(* Logix 5000 project; controller OWF Emulate 5570 rev 30.12; software revision 30.00 *) (continued)
   	OWF_Key[222,1]:=1243582292;
   	OWF_Key[222,2]:=1667078718;
   	OWF_Key[222,3]:=820047921;
   	OWF_Key[222,4]:=2100818839;
   	OWF_Key[222,5]:=54664303;
   	OWF_Key[222,6]:=832390246;
   	OWF_Key[222,7]:=1025838178;
   	OWF_Key[222,8]:=2108609866;
   	OWF_Key[223,0]:=1550121582;
   	OWF_Key[223,1]:=901840231;
   	OWF_Key[223,2]:=845237975;
   	OWF_Key[223,3]:=1737038115;
   	OWF_Key[223,4]:=250371253;
   	OWF_Key[223,5]:=841400060;
   	OWF_Key[223,6]:=633458828;
   	OWF_Key[223,7]:=1234192716;
   	OWF_Key[223,8]:=1638825880;
   	OWF_Key[224,0]:=1100202784;
   	OWF_Key[224,1]:=1268618722;
   	OWF_Key[224,2]:=1328247563;
   	OWF_Key[224,3]:=315030373;
   	OWF_Key[224,4]:=17465755;
   	OWF_Key[224,5]:=1489898403;
   	OWF_Key[224,6]:=1369322265;
   	OWF_Key[224,7]:=2029664960;
   	OWF_Key[224,8]:=1183192871;
   	OWF_Key[225,0]:=1841076227;
   	OWF_Key[225,1]:=1387440943;
   	OWF_Key[225,2]:=94964990;
   	OWF_Key[225,3]:=374620338;
   	OWF_Key[225,4]:=198656364;
   	OWF_Key[225,5]:=451329169;
   	OWF_Key[225,6]:=1040984125;
   	OWF_Key[225,7]:=421870535;
   	OWF_Key[225,8]:=1711294224;
   	OWF_Key[226,0]:=908174588;
   	OWF_Key[226,1]:=915800259;
   	OWF_Key[226,2]:=1938292132;
   	OWF_Key[226,3]:=1295597437;
   	OWF_Key[226,4]:=543239841;
   	OWF_Key[226,5]:=543313500;
   	OWF_Key[226,6]:=1320318736;
   	OWF_Key[226,7]:=1310833438;
   	OWF_Key[226,8]:=1604355088;
   	OWF_Key[227,0]:=1963899269;
   	OWF_Key[227,1]:=1680451206;
   	OWF_Key[227,2]:=236776837;
   	OWF_Key[227,3]:=1960573892;
   	OWF_Key[227,4]:=2100303206;
   	OWF_Key[227,5]:=407078522;
   	OWF_Key[227,6]:=949933681;
   	OWF_Key[227,7]:=279399557;
   	OWF_Key[227,8]:=510170757;
   	OWF_Key[228,0]:=407858862;
   	OWF_Key[228,1]:=1041535109;
   	OWF_Key[228,2]:=75109540;
   	OWF_Key[228,3]:=341906229;
   	OWF_Key[228,4]:=1034027359;
   	OWF_Key[228,5]:=899760418;
   	OWF_Key[228,6]:=1758227630;
   	OWF_Key[228,7]:=2129936455;
   	OWF_Key[228,8]:=914417718;
   	OWF_Key[229,0]:=649884288;
   	OWF_Key[229,1]:=926898577;
   	OWF_Key[229,2]:=189532880;
   	OWF_Key[229,3]:=262049990;
   	OWF_Key[229,4]:=1071612823;
   	OWF_Key[229,5]:=63876222;
   	OWF_Key[229,6]:=581163575;
   	OWF_Key[229,7]:=537068257;
   	OWF_Key[229,8]:=266266259;
   	OWF_Key[230,0]:=2037870100;
   	OWF_Key[230,1]:=953538015;
   	OWF_Key[230,2]:=1215162513;
   	OWF_Key[230,3]:=1204636685;
   	OWF_Key[230,4]:=1759636210;
   	OWF_Key[230,5]:=1064005198;
   	OWF_Key[230,6]:=183113685;
   	OWF_Key[230,7]:=732180321;
   	OWF_Key[230,8]:=755593610;
   	OWF_Key[231,0]:=210769631;
   	OWF_Key[231,1]:=171144649;
   	OWF_Key[231,2]:=453217172;
   	OWF_Key[231,3]:=1410128994;
   	OWF_Key[231,4]:=1742068836;
   	OWF_Key[231,5]:=1433828688;
   	OWF_Key[231,6]:=1733251173;
   	OWF_Key[231,7]:=175140488;
   	OWF_Key[231,8]:=1694955713;
   	OWF_Key[232,0]:=754935092;
   	OWF_Key[232,1]:=1561205565;
   	OWF_Key[232,2]:=1437601257;
   	OWF_Key[232,3]:=1566278877;
   	OWF_Key[232,4]:=592341060;
   	OWF_Key[232,5]:=296146351;
   	OWF_Key[232,6]:=1009239711;
   	OWF_Key[232,7]:=1066032517;
   	OWF_Key[232,8]:=1401251796;
   	OWF_Key[233,0]:=2014784236;
   	OWF_Key[233,1]:=210556685;
   	OWF_Key[233,2]:=603004710;
   	OWF_Key[233,3]:=2050599314;
   	OWF_Key[233,4]:=1831548063;
   	OWF_Key[233,5]:=1680385195;
   	OWF_Key[233,6]:=46017568;
   	OWF_Key[233,7]:=806626447;
   	OWF_Key[233,8]:=429224258;
   	OWF_Key[234,0]:=102806102;
   	OWF_Key[234,1]:=1249179697;
   	OWF_Key[234,2]:=1376509434;
   	OWF_Key[234,3]:=519963743;
   	OWF_Key[234,4]:=1266509533;
   	OWF_Key[234,5]:=1500035180;
   	OWF_Key[234,6]:=1362314000;
   	OWF_Key[234,7]:=270021354;
   	OWF_Key[234,8]:=1980281736;
   	OWF_Key[235,0]:=1108202131;
   	OWF_Key[235,1]:=364018967;
   	OWF_Key[235,2]:=2002036400;
   	OWF_Key[235,3]:=287661169;
   	OWF_Key[235,4]:=163785897;
   	OWF_Key[235,5]:=1093258499;
   	OWF_Key[235,6]:=595570472;
   	OWF_Key[235,7]:=1298504233;
   	OWF_Key[235,8]:=1061993871;
   	OWF_Key[236,0]:=754930847;
   	OWF_Key[236,1]:=1771686064;
   	OWF_Key[236,2]:=1612117580;
   	OWF_Key[236,3]:=78834364;
   	OWF_Key[236,4]:=2112379245;
   	OWF_Key[236,5]:=685652796;
   	OWF_Key[236,6]:=361207730;
   	OWF_Key[236,7]:=134397244;
   	OWF_Key[236,8]:=1371411455;
   	OWF_Key[237,0]:=2093988696;
   	OWF_Key[237,1]:=1048911586;
   	OWF_Key[237,2]:=832606970;
   	OWF_Key[237,3]:=1492019873;
   	OWF_Key[237,4]:=1423376112;
   	OWF_Key[237,5]:=38580303;
   	OWF_Key[237,6]:=868576798;
   	OWF_Key[237,7]:=1397461282;
   	OWF_Key[237,8]:=960767099;
   	OWF_Key[238,0]:=1250673699;
   	OWF_Key[238,1]:=1617635287;
   	OWF_Key[238,2]:=470819108;
   	OWF_Key[238,3]:=959348674;
   	OWF_Key[238,4]:=1001458249;
   	OWF_Key[238,5]:=1747882864;
   	OWF_Key[238,6]:=1322152057;
   	OWF_Key[238,7]:=679295127;
   	OWF_Key[238,8]:=1876556191;
   	OWF_Key[239,0]:=36757702;
   	OWF_Key[239,1]:=1049474760;
   	OWF_Key[239,2]:=1824982906;
   	OWF_Key[239,3]:=2096596441;
   	OWF_Key[239,4]:=1687250299;
   	OWF_Key[239,5]:=1833823020;
   	OWF_Key[239,6]:=686257311;
   	OWF_Key[239,7]:=1367821520;
   	OWF_Key[239,8]:=1928845366;
   	OWF_Key[240,0]:=1169899109;
   	OWF_Key[240,1]:=1726445489;
   	OWF_Key[240,2]:=50823841;
   	OWF_Key[240,3]:=908212678;
   	OWF_Key[240,4]:=1158043459;
   	OWF_Key[240,5]:=98435470;
   	OWF_Key[240,6]:=590448747;
   	OWF_Key[240,7]:=610552049;
   	OWF_Key[240,8]:=614864981;
   	OWF_Key[241,0]:=1140035422;
   	OWF_Key[241,1]:=1630773789;
   	OWF_Key[241,2]:=1291895646;
   	OWF_Key[241,3]:=1981816599;
   	OWF_Key[241,4]:=1262307061;
   	OWF_Key[241,5]:=122395708;
   	OWF_Key[241,6]:=817314502;
   	OWF_Key[241,7]:=519742265;
   	OWF_Key[241,8]:=444078296;
   	OWF_Key[242,0]:=821076122;
   	OWF_Key[242,1]:=205468863;
   	OWF_Key[242,2]:=1709938843;
   	OWF_Key[242,3]:=250210989;
   	OWF_Key[242,4]:=725159142;
   	OWF_Key[242,5]:=1933164860;
   	OWF_Key[242,6]:=1311047082;
   	OWF_Key[242,7]:=79103381;
   	OWF_Key[242,8]:=1836791040;
   	OWF_Key[243,0]:=604446577;
   	OWF_Key[243,1]:=1973034181;
   	OWF_Key[243,2]:=1229878013;
   	OWF_Key[243,3]:=313423778;
   	OWF_Key[243,4]:=1453913733;
   	OWF_Key[243,5]:=136665972;
   	OWF_Key[243,6]:=1095058148;
   	OWF_Key[243,7]:=1245422719;
   	OWF_Key[243,8]:=1645758259;
   	OWF_Key[244,0]:=1415797906;
   	OWF_Key[244,1]:=1697757892;
   	OWF_Key[244,2]:=759890877;
   	OWF_Key[244,3]:=24103685;
   	OWF_Key[244,4]:=1909169002;
   	OWF_Key[244,5]:=922218833;
   	OWF_Key[244,6]:=1165355415;
   	OWF_Key[244,7]:=1904308279;
   	OWF_Key[244,8]:=638820940;
   	OWF_Key[245,0]:=301200093;
   	OWF_Key[245,1]:=1314891726;
   	OWF_Key[245,2]:=692781419;
   	OWF_Key[245,3]:=2023891545;
   	OWF_Key[245,4]:=746992191;
   	OWF_Key[245,5]:=769066877;
   	OWF_Key[245,6]:=670754800;
   	OWF_Key[245,7]:=1544280754;
   	OWF_Key[245,8]:=399959487;
   	OWF_Key[246,0]:=74045861;
   	OWF_Key[246,1]:=58012275;
   	OWF_Key[246,2]:=767892604;
   	OWF_Key[246,3]:=1587247299;
   	OWF_Key[246,4]:=914262113;
   	OWF_Key[246,5]:=759782505;
   	OWF_Key[246,6]:=1121680670;
   	OWF_Key[246,7]:=1483043544;
   	OWF_Key[246,8]:=578023515;
   	OWF_Key[247,0]:=468948122;
   	OWF_Key[247,1]:=323506121;
   	OWF_Key[247,2]:=1230071484;
   	OWF_Key[247,3]:=748609841;
   	OWF_Key[247,4]:=177788530;
   	OWF_Key[247,5]:=618957179;
   	OWF_Key[247,6]:=1569691208;
   	OWF_Key[247,7]:=534187793;
   	OWF_Key[247,8]:=15501750;
   	OWF_Key[248,0]:=1850366820;
   	OWF_Key[248,1]:=1406619300;
   	OWF_Key[248,2]:=1237604397;
   	OWF_Key[248,3]:=1081902870;
   	OWF_Key[248,4]:=1641259906;
   	OWF_Key[248,5]:=125727550;
   	OWF_Key[248,6]:=1749051731;
   	OWF_Key[248,7]:=1967031533;
   	OWF_Key[248,8]:=1220540139;
   	OWF_Key[249,0]:=100619500;
   	OWF_Key[249,1]:=1511118985;
   	OWF_Key[249,2]:=106143349;
   	OWF_Key[249,3]:=710065616;
   	OWF_Key[249,4]:=1830124358;
   	OWF_Key[249,5]:=985511526;
   	OWF_Key[249,6]:=2059823479;
   	OWF_Key[249,7]:=1691454625;
   	OWF_Key[249,8]:=966899445;
   	OWF_Key[250,0]:=664287990;
   	OWF_Key[250,1]:=1886466319;
   	OWF_Key[250,2]:=956844688;
   	OWF_Key[250,3]:=1061940606;
   	OWF_Key[250,4]:=1037885088;
   	OWF_Key[250,5]:=311608117;
   	OWF_Key[250,6]:=2003988095;
   	OWF_Key[250,7]:=1878351249;
   	OWF_Key[250,8]:=811092189;
   	OWF_Key[251,0]:=27430717;
   	OWF_Key[251,1]:=141278967;
   	OWF_Key[251,2]:=1720155622;
   	OWF_Key[251,3]:=737827649;
   	OWF_Key[251,4]:=238939021;
   	OWF_Key[251,5]:=538882310;
   	OWF_Key[251,6]:=1366554664;
   	OWF_Key[251,7]:=1186610005;
   	OWF_Key[251,8]:=817820658;
   	OWF_Key[252,0]:=1867493799;
   	OWF_Key[252,1]:=1604329457;
   	OWF_Key[252,2]:=238680985;
   	OWF_Key[252,3]:=1920811059;
   	OWF_Key[252,4]:=748517017;
   	OWF_Key[252,5]:=969165835;
   	OWF_Key[252,6]:=1811752884;
   	OWF_Key[252,7]:=1156638675;
   	OWF_Key[252,8]:=287327869;
   	OWF_Key[253,0]:=327334567;
   	OWF_Key[253,1]:=938516870;
   	OWF_Key[253,2]:=1209234380;
   	OWF_Key[253,3]:=1945410057;
   	OWF_Key[253,4]:=1246767444;
   	OWF_Key[253,5]:=1539463706;
   	OWF_Key[253,6]:=1541419964;
   	OWF_Key[253,7]:=675055296;
   	OWF_Key[253,8]:=1234478343;
   	OWF_Key[254,0]:=220047547;
   	OWF_Key[254,1]:=1437897813;
   	OWF_Key[254,2]:=1852012355;
   	OWF_Key[254,3]:=1583044272;
   	OWF_Key[254,4]:=228664887;
   	OWF_Key[254,5]:=1600113842;
   	OWF_Key[254,6]:=98868957;
   	OWF_Key[254,7]:=899477217;
   	OWF_Key[254,8]:=2080520664;
   	OWF_Key[255,0]:=221865779;
   	OWF_Key[255,1]:=729341680;
   	OWF_Key[255,2]:=1616592850;
   	OWF_Key[255,3]:=1543315716;
   	OWF_Key[255,4]:=1981504727;
   	OWF_Key[255,5]:=1919924645;
   	OWF_Key[255,6]:=400471940;
   	OWF_Key[255,7]:=337852422;
   	OWF_Key[255,8]:=128006188;
   End_If;
   If OWF_Ver > 0 Then
   	OWF_Key[0,9]:=565857393;
   	OWF_Key[0,10]:=1292544462;
   	OWF_Key[0,11]:=880397583;
   	OWF_Key[0,12]:=526971504;
   	OWF_Key[1,9]:=136125333;
   	OWF_Key[1,10]:=772079857;
   	OWF_Key[1,11]:=262884596;
   	OWF_Key[1,12]:=1285068215;
   	OWF_Key[2,9]:=1935405231;
   	OWF_Key[2,10]:=1279162383;
   	OWF_Key[2,11]:=316222445;
   	OWF_Key[2,12]:=52577038;
   	OWF_Key[3,9]:=462041571;
   	OWF_Key[3,10]:=944242743;
   	OWF_Key[3,11]:=1789622395;
   	OWF_Key[3,12]:=1944538496;
   	OWF_Key[4,9]:=1444514190;
   	OWF_Key[4,10]:=1887503071;
   	OWF_Key[4,11]:=4758697;
   	OWF_Key[4,12]:=1055291277;
   	OWF_Key[5,9]:=1069465770;
   	OWF_Key[5,10]:=956524197;
   	OWF_Key[5,11]:=772219220;
   	OWF_Key[5,12]:=1564477108;
   	OWF_Key[6,9]:=527419559;
   	OWF_Key[6,10]:=2004204950;
   	OWF_Key[6,11]:=28698575;
   	OWF_Key[6,12]:=214680673;
   	OWF_Key[7,9]:=1681234259;
   	OWF_Key[7,10]:=580130361;
   	OWF_Key[7,11]:=1396051131;
   	OWF_Key[7,12]:=1471817513;
   	OWF_Key[8,9]:=445296913;
   	OWF_Key[8,10]:=1852602746;
   	OWF_Key[8,11]:=663900175;
   	OWF_Key[8,12]:=480645843;
   	OWF_Key[9,9]:=911927794;
   	OWF_Key[9,10]:=2147066014;
   	OWF_Key[9,11]:=1002765035;
   	OWF_Key[9,12]:=1677182369;
   	OWF_Key[10,9]:=449913502;
   	OWF_Key[10,10]:=1451210493;
   	OWF_Key[10,11]:=1560758298;
   	OWF_Key[10,12]:=1653399395;
   	OWF_Key[11,9]:=336562059;
   	OWF_Key[11,10]:=460160972;
   	OWF_Key[11,11]:=267446441;
   	OWF_Key[11,12]:=1872890613;
   	OWF_Key[12,9]:=1991253080;
   	OWF_Key[12,10]:=326769400;
   	OWF_Key[12,11]:=1075259094;
   	OWF_Key[12,12]:=39472927;
   	OWF_Key[13,9]:=1611056956;
   	OWF_Key[13,10]:=109533992;
   	OWF_Key[13,11]:=1225494993;
   	OWF_Key[13,12]:=859906139;
   	OWF_Key[14,9]:=1244611515;
   	OWF_Key[14,10]:=442554456;
   	OWF_Key[14,11]:=1104886967;
   	OWF_Key[14,12]:=726142142;
   	OWF_Key[15,9]:=640501099;
   	OWF_Key[15,10]:=475719934;
   	OWF_Key[15,11]:=25495759;
   	OWF_Key[15,12]:=780644316;
   	OWF_Key[16,9]:=1277928375;
   	OWF_Key[16,10]:=1138754243;
   	OWF_Key[16,11]:=426325284;
   	OWF_Key[16,12]:=962841358;
   	OWF_Key[17,9]:=81801666;
   	OWF_Key[17,10]:=702205204;
   	OWF_Key[17,11]:=1750566476;
   	OWF_Key[17,12]:=658348297;
   	OWF_Key[18,9]:=1606390434;
   	OWF_Key[18,10]:=553184116;
   	OWF_Key[18,11]:=92452548;
   	OWF_Key[18,12]:=544582854;
   	OWF_Key[19,9]:=2075044410;
   	OWF_Key[19,10]:=955756930;
   	OWF_Key[19,11]:=623976828;
   	OWF_Key[19,12]:=135043920;
   	OWF_Key[20,9]:=755768755;
   	OWF_Key[20,10]:=195409842;
   	OWF_Key[20,11]:=484943474;
   	OWF_Key[20,12]:=1966535273;
   	OWF_Key[21,9]:=1524021832;
   	OWF_Key[21,10]:=553649431;
   	OWF_Key[21,11]:=1634240438;
   	OWF_Key[21,12]:=233480851;
   	OWF_Key[22,9]:=2044449579;
   	OWF_Key[22,10]:=1409976464;
   	OWF_Key[22,11]:=261784018;
   	OWF_Key[22,12]:=769448317;
   	OWF_Key[23,9]:=995187060;
   	OWF_Key[23,10]:=422401363;
   	OWF_Key[23,11]:=108903649;
   	OWF_Key[23,12]:=2052854235;
   	OWF_Key[24,9]:=848694715;
   	OWF_Key[24,10]:=1665199255;
   	OWF_Key[24,11]:=2100798558;
   	OWF_Key[24,12]:=1683952239;
   	OWF_Key[25,9]:=743358321;
   	OWF_Key[25,10]:=1278338921;
   	OWF_Key[25,11]:=317357624;
   	OWF_Key[25,12]:=42763409;
   	OWF_Key[26,9]:=1269606561;
   	OWF_Key[26,10]:=791897924;
   	OWF_Key[26,11]:=604881525;
   	OWF_Key[26,12]:=1224898459;
   	OWF_Key[27,9]:=1927567431;
   	OWF_Key[27,10]:=375986974;
   	OWF_Key[27,11]:=1705499705;
   	OWF_Key[27,12]:=668949563;
   	OWF_Key[28,9]:=1045167080;
   	OWF_Key[28,10]:=41953216;
   	OWF_Key[28,11]:=1054662341;
   	OWF_Key[28,12]:=1395343957;
   	OWF_Key[29,9]:=865673428;
   	OWF_Key[29,10]:=2145157796;
   	OWF_Key[29,11]:=1458425611;
   	OWF_Key[29,12]:=205894898;
   	OWF_Key[30,9]:=731876933;
   	OWF_Key[30,10]:=1676387747;
   	OWF_Key[30,11]:=945162642;
   	OWF_Key[30,12]:=331348069;
   	OWF_Key[31,9]:=280733610;
   	OWF_Key[31,10]:=440691357;
   	OWF_Key[31,11]:=919012913;
   	OWF_Key[31,12]:=1726573128;
   	OWF_Key[32,9]:=1387391898;
   	OWF_Key[32,10]:=1975692002;
   	OWF_Key[32,11]:=1709706860;
   	OWF_Key[32,12]:=763727752;
   	OWF_Key[33,9]:=752730332;
   	OWF_Key[33,10]:=1724856462;
   	OWF_Key[33,11]:=654259641;
   	OWF_Key[33,12]:=1291634161;
   	OWF_Key[34,9]:=547087700;
   	OWF_Key[34,10]:=1022930882;
   	OWF_Key[34,11]:=409869923;
   	OWF_Key[34,12]:=1072376958;
   	OWF_Key[35,9]:=1977060651;
   	OWF_Key[35,10]:=765565508;
   	OWF_Key[35,11]:=2104021265;
   	OWF_Key[35,12]:=1906749018;
   	OWF_Key[36,9]:=1927629184;
   	OWF_Key[36,10]:=1689263679;
   	OWF_Key[36,11]:=1705229799;
   	OWF_Key[36,12]:=767108731;
   	OWF_Key[37,9]:=1051908007;
   	OWF_Key[37,10]:=737157349;
   	OWF_Key[37,11]:=1462539168;
   	OWF_Key[37,12]:=954814956;
   	OWF_Key[38,9]:=215452186;
   	OWF_Key[38,10]:=741757339;
   	OWF_Key[38,11]:=988659375;
   	OWF_Key[38,12]:=1743432283;
   	OWF_Key[39,9]:=1418135291;
   	OWF_Key[39,10]:=1958452124;
   	OWF_Key[39,11]:=1028640656;
   	OWF_Key[39,12]:=1067663543;
   	OWF_Key[40,9]:=1684938390;
   	OWF_Key[40,10]:=651300804;
   	OWF_Key[40,11]:=515025545;
   	OWF_Key[40,12]:=1116941873;
   	OWF_Key[41,9]:=1635688259;
   	OWF_Key[41,10]:=1065432902;
   	OWF_Key[41,11]:=1719788305;
   	OWF_Key[41,12]:=626834989;
   	OWF_Key[42,9]:=1581635246;
   	OWF_Key[42,10]:=1478705635;
   	OWF_Key[42,11]:=2022105722;
   	OWF_Key[42,12]:=1757031333;
   	OWF_Key[43,9]:=2019000851;
   	OWF_Key[43,10]:=552604579;
   	OWF_Key[43,11]:=346246408;
   	OWF_Key[43,12]:=714285990;
   	OWF_Key[44,9]:=49056678;
   	OWF_Key[44,10]:=1632958150;
   	OWF_Key[44,11]:=190550872;
   	OWF_Key[44,12]:=478927043;
   	OWF_Key[45,9]:=35435192;
   	OWF_Key[45,10]:=516712311;
   	OWF_Key[45,11]:=257768150;
   	OWF_Key[45,12]:=193871838;
   	OWF_Key[46,9]:=446657733;
   	OWF_Key[46,10]:=1362936296;
   	OWF_Key[46,11]:=936691800;
   	OWF_Key[46,12]:=1446652431;
   	OWF_Key[47,9]:=174593183;
   	OWF_Key[47,10]:=264816060;
   	OWF_Key[47,11]:=239257452;
   	OWF_Key[47,12]:=1557535775;
   	OWF_Key[48,9]:=23082539;
   	OWF_Key[48,10]:=1885756789;
   	OWF_Key[48,11]:=2139584242;
   	OWF_Key[48,12]:=567181888;
   	OWF_Key[49,9]:=59195043;
   	OWF_Key[49,10]:=832903498;
   	OWF_Key[49,11]:=115146831;
   	OWF_Key[49,12]:=1133120569;
   	OWF_Key[50,9]:=1265526322;
   	OWF_Key[50,10]:=114687092;
   	OWF_Key[50,11]:=1570753334;
   	OWF_Key[50,12]:=1848310255;
   	OWF_Key[51,9]:=2088557685;
   	OWF_Key[51,10]:=1083470336;
   	OWF_Key[51,11]:=952144566;
   	OWF_Key[51,12]:=1526744395;
   	OWF_Key[52,9]:=778318022;
   	OWF_Key[52,10]:=415429748;
   	OWF_Key[52,11]:=1695256824;
   	OWF_Key[52,12]:=677148294;
   	OWF_Key[53,9]:=968528232;
   	OWF_Key[53,10]:=1557455946;
   	OWF_Key[53,11]:=1203553962;
   	OWF_Key[53,12]:=960333575;
   	OWF_Key[54,9]:=511483668;
   	OWF_Key[54,10]:=2051447889;
   	OWF_Key[54,11]:=452797653;
   	OWF_Key[54,12]:=929742413;
   	OWF_Key[55,9]:=1860951280;
   	OWF_Key[55,10]:=1206370150;
   	OWF_Key[55,11]:=840015040;
   	OWF_Key[55,12]:=2012424497;
   	OWF_Key[56,9]:=1960686173;
   	OWF_Key[56,10]:=292188386;
   	OWF_Key[56,11]:=1295478345;
   	OWF_Key[56,12]:=134139962;
   	OWF_Key[57,9]:=1725868720;
   	OWF_Key[57,10]:=1022760847;
   	OWF_Key[57,11]:=1266867308;
   	OWF_Key[57,12]:=1518331712;
   	OWF_Key[58,9]:=1287898341;
   	OWF_Key[58,10]:=1112687552;
   	OWF_Key[58,11]:=1981827060;
   	OWF_Key[58,12]:=1854707709;
   	OWF_Key[59,9]:=1826891165;
   	OWF_Key[59,10]:=1690535487;
   	OWF_Key[59,11]:=1854035272;
   	OWF_Key[59,12]:=2145802432;
   	OWF_Key[60,9]:=2116204488;
   	OWF_Key[60,10]:=598097181;
   	OWF_Key[60,11]:=1722801485;
   	OWF_Key[60,12]:=1928154342;
   	OWF_Key[61,9]:=290230891;
   	OWF_Key[61,10]:=139306183;
   	OWF_Key[61,11]:=1302319781;
   	OWF_Key[61,12]:=1778862980;
   	OWF_Key[62,9]:=1398911657;
   	OWF_Key[62,10]:=795615750;
   	OWF_Key[62,11]:=1649806734;
   	OWF_Key[62,12]:=730523144;
   	OWF_Key[63,9]:=509322045;
   	OWF_Key[63,10]:=1394809523;
   	OWF_Key[63,11]:=1242281877;
   	OWF_Key[63,12]:=1337104856;
   	OWF_Key[64,9]:=520494279;
   	OWF_Key[64,10]:=1407862991;
   	OWF_Key[64,11]:=601636969;
   	OWF_Key[64,12]:=984487298;
   	OWF_Key[65,9]:=2040473319;
   	OWF_Key[65,10]:=1825501221;
   	OWF_Key[65,11]:=719189220;
   	OWF_Key[65,12]:=1705052589;
   	OWF_Key[66,9]:=614095249;
   	OWF_Key[66,10]:=1060379412;
   	OWF_Key[66,11]:=818790030;
   	OWF_Key[66,12]:=2082342074;
   	OWF_Key[67,9]:=379359286;
   	OWF_Key[67,10]:=625025710;
   	OWF_Key[67,11]:=581201342;
   	OWF_Key[67,12]:=1291639086;
   	OWF_Key[68,9]:=2034139144;
   	OWF_Key[68,10]:=1775077551;
   	OWF_Key[68,11]:=1149406496;
   	OWF_Key[68,12]:=487904912;
   	OWF_Key[69,9]:=1508683351;
   	OWF_Key[69,10]:=1277536059;
   	OWF_Key[69,11]:=967303233;
   	OWF_Key[69,12]:=1006071908;
   	OWF_Key[70,9]:=1502345175;
   	OWF_Key[70,10]:=682860158;
   	OWF_Key[70,11]:=784529015;
   	OWF_Key[70,12]:=561765580;
   	OWF_Key[71,9]:=1817547816;
   	OWF_Key[71,10]:=1507525691;
   	OWF_Key[71,11]:=255509082;
   	OWF_Key[71,12]:=1551741993;
   	OWF_Key[72,9]:=629806228;
   	OWF_Key[72,10]:=571635577;
   	OWF_Key[72,11]:=1224031942;
   	OWF_Key[72,12]:=181619567;
   	OWF_Key[73,9]:=1469724584;
   	OWF_Key[73,10]:=594076044;
   	OWF_Key[73,11]:=1411066369;
   	OWF_Key[73,12]:=550406167;
   	OWF_Key[74,9]:=1331101818;
   	OWF_Key[74,10]:=339372374;
   	OWF_Key[74,11]:=988614620;
   	OWF_Key[74,12]:=116767437;
   	OWF_Key[75,9]:=158649017;
   	OWF_Key[75,10]:=782737333;
   	OWF_Key[75,11]:=530692638;
   	OWF_Key[75,12]:=808012468;
   	OWF_Key[76,9]:=1154486896;
   	OWF_Key[76,10]:=405198090;
   	OWF_Key[76,11]:=542834227;
   	OWF_Key[76,12]:=1280285599;
   	OWF_Key[77,9]:=1474337535;
   	OWF_Key[77,10]:=1523725108;
   	OWF_Key[77,11]:=2145251389;
   	OWF_Key[77,12]:=1246513416;
   	OWF_Key[78,9]:=1162275216;
   	OWF_Key[78,10]:=961731882;
   	OWF_Key[78,11]:=1909965356;
   	OWF_Key[78,12]:=1970279923;
   	OWF_Key[79,9]:=812018256;
   	OWF_Key[79,10]:=59709690;
   	OWF_Key[79,11]:=1481776184;
   	OWF_Key[79,12]:=355946496;
   	OWF_Key[80,9]:=1668122452;
   	OWF_Key[80,10]:=1498872612;
   	OWF_Key[80,11]:=1612349490;
   	OWF_Key[80,12]:=1851589051;
   	OWF_Key[81,9]:=1599256517;
   	OWF_Key[81,10]:=912097274;
   	OWF_Key[81,11]:=679219195;
   	OWF_Key[81,12]:=744308687;
   	OWF_Key[82,9]:=1233315062;
   	OWF_Key[82,10]:=2129485434;
   	OWF_Key[82,11]:=1977811005;
   	OWF_Key[82,12]:=194772472;
   	OWF_Key[83,9]:=452177585;
   	OWF_Key[83,10]:=2103129384;
   	OWF_Key[83,11]:=1881046621;
   	OWF_Key[83,12]:=262049613;
   	OWF_Key[84,9]:=591161416;
   	OWF_Key[84,10]:=2029877352;
   	OWF_Key[84,11]:=47581452;
   	OWF_Key[84,12]:=926767567;
   	OWF_Key[85,9]:=1823347902;
   	OWF_Key[85,10]:=499556028;
   	OWF_Key[85,11]:=1207806672;
   	OWF_Key[85,12]:=1702523720;
   	OWF_Key[86,9]:=48595898;
   	OWF_Key[86,10]:=872429374;
   	OWF_Key[86,11]:=66297910;
   	OWF_Key[86,12]:=1790557355;
   	OWF_Key[87,9]:=403726996;
   	OWF_Key[87,10]:=1458912687;
   	OWF_Key[87,11]:=24431334;
   	OWF_Key[87,12]:=1173086986;
   	OWF_Key[88,9]:=39924540;
   	OWF_Key[88,10]:=1496951722;
   	OWF_Key[88,11]:=1856630873;
   	OWF_Key[88,12]:=1127631222;
   	OWF_Key[89,9]:=669788712;
   	OWF_Key[89,10]:=1130692876;
   	OWF_Key[89,11]:=1518579924;
   	OWF_Key[89,12]:=1718912249;
   	OWF_Key[90,9]:=978095313;
   	OWF_Key[90,10]:=1619784712;
   	OWF_Key[90,11]:=1680494857;
   	OWF_Key[90,12]:=1794312175;
   	OWF_Key[91,9]:=322164715;
   	OWF_Key[91,10]:=511187759;
   	OWF_Key[91,11]:=554109920;
   	OWF_Key[91,12]:=1832701750;
   	OWF_Key[92,9]:=1289671026;
   	OWF_Key[92,10]:=1720186424;
   	OWF_Key[92,11]:=762336602;
   	OWF_Key[92,12]:=594253437;
   	OWF_Key[93,9]:=754238063;
   	OWF_Key[93,10]:=101706781;
   	OWF_Key[93,11]:=552270309;
   	OWF_Key[93,12]:=470087240;
   	OWF_Key[94,9]:=1836214779;
   	OWF_Key[94,10]:=1972536857;
   	OWF_Key[94,11]:=732394613;
   	OWF_Key[94,12]:=550096746;
   	OWF_Key[95,9]:=1681612441;
   	OWF_Key[95,10]:=1464436621;
   	OWF_Key[95,11]:=851826791;
   	OWF_Key[95,12]:=1584332130;
   	OWF_Key[96,9]:=1811817677;
   	OWF_Key[96,10]:=1389118238;
   	OWF_Key[96,11]:=1984755030;
   	OWF_Key[96,12]:=1486487521;
   	OWF_Key[97,9]:=1937715549;
   	OWF_Key[97,10]:=455909523;
   	OWF_Key[97,11]:=693528960;
   	OWF_Key[97,12]:=484997079;
   	OWF_Key[98,9]:=593189665;
   	OWF_Key[98,10]:=716154395;
   	OWF_Key[98,11]:=634179513;
   	OWF_Key[98,12]:=1431023684;
   	OWF_Key[99,9]:=1303410798;
   	OWF_Key[99,10]:=1929791531;
   	OWF_Key[99,11]:=1153562302;
   	OWF_Key[99,12]:=983138799;
   	OWF_Key[100,9]:=1831590352;
   	OWF_Key[100,10]:=626802806;
   	OWF_Key[100,11]:=950067436;
   	OWF_Key[100,12]:=1058805733;
   	OWF_Key[101,9]:=254358295;
   	OWF_Key[101,10]:=1733530591;
   	OWF_Key[101,11]:=1763235204;
   	OWF_Key[101,12]:=3204015;
   	OWF_Key[102,9]:=1824511525;
   	OWF_Key[102,10]:=1242921701;
   	OWF_Key[102,11]:=1037008908;
   	OWF_Key[102,12]:=1819226588;
   	OWF_Key[103,9]:=375657977;
   	OWF_Key[103,10]:=434997384;
   	OWF_Key[103,11]:=1632163593;
   	OWF_Key[103,12]:=1224085853;
   	OWF_Key[104,9]:=834825299;
   	OWF_Key[104,10]:=1757006557;
   	OWF_Key[104,11]:=1725971178;
   	OWF_Key[104,12]:=758876662;
   	OWF_Key[105,9]:=1632620875;
   	OWF_Key[105,10]:=164276743;
   	OWF_Key[105,11]:=1757534671;
   	OWF_Key[105,12]:=49011059;
   	OWF_Key[106,9]:=1924183141;
   	OWF_Key[106,10]:=1377114833;
   	OWF_Key[106,11]:=1520087306;
   	OWF_Key[106,12]:=403124570;
   	OWF_Key[107,9]:=1476158981;
   	OWF_Key[107,10]:=472928532;
   	OWF_Key[107,11]:=1763552980;
   	OWF_Key[107,12]:=2082172463;
   	OWF_Key[108,9]:=1432733723;
   	OWF_Key[108,10]:=1041871619;
   	OWF_Key[108,11]:=848827879;
   	OWF_Key[108,12]:=761199130;
   	OWF_Key[109,9]:=1437046258;
   	OWF_Key[109,10]:=1857419035;
   	OWF_Key[109,11]:=1735010683;
   	OWF_Key[109,12]:=944312109;
   	OWF_Key[110,9]:=1543386268;
   	OWF_Key[110,10]:=1134207558;
   	OWF_Key[110,11]:=2101947387;
   	OWF_Key[110,12]:=1169923182;
   	OWF_Key[111,9]:=194570507;
   	OWF_Key[111,10]:=717684516;
   	OWF_Key[111,11]:=2027079632;
   	OWF_Key[111,12]:=281935625;
   	OWF_Key[112,9]:=1723553691;
   	OWF_Key[112,10]:=820691500;
   	OWF_Key[112,11]:=1726230371;
   	OWF_Key[112,12]:=2140435056;
   	OWF_Key[113,9]:=422933751;
   	OWF_Key[113,10]:=1361381455;
   	OWF_Key[113,11]:=503450599;
   	OWF_Key[113,12]:=176022433;
   	OWF_Key[114,9]:=947522075;
   	OWF_Key[114,10]:=2041241092;
   	OWF_Key[114,11]:=354278848;
   	OWF_Key[114,12]:=1134259119;
   	OWF_Key[115,9]:=534251520;
   	OWF_Key[115,10]:=1093413069;
   	OWF_Key[115,11]:=1469054204;
   	OWF_Key[115,12]:=1011873089;
   	OWF_Key[116,9]:=2110878619;
   	OWF_Key[116,10]:=391290202;
   	OWF_Key[116,11]:=2077826702;
   	OWF_Key[116,12]:=1896888156;
   	OWF_Key[117,9]:=890737217;
   	OWF_Key[117,10]:=1056381272;
   	OWF_Key[117,11]:=1732884181;
   	OWF_Key[117,12]:=948255347;
   	OWF_Key[118,9]:=2140498942;
   	OWF_Key[118,10]:=1215633590;
   	OWF_Key[118,11]:=724300285;
   	OWF_Key[118,12]:=309190363;
   	OWF_Key[119,9]:=301015591;
   	OWF_Key[119,10]:=1841175439;
   	OWF_Key[119,11]:=1489747792;
   	OWF_Key[119,12]:=990396034;
   	OWF_Key[120,9]:=1029365379;
   	OWF_Key[120,10]:=685059449;
   	OWF_Key[120,11]:=561217780;
   	OWF_Key[120,12]:=908603653;
   	OWF_Key[121,9]:=651112791;
   	OWF_Key[121,10]:=1007517130;
   	OWF_Key[121,11]:=430229034;
   	OWF_Key[121,12]:=741552407;
   	OWF_Key[122,9]:=205699509;
   	OWF_Key[122,10]:=1591187346;
   	OWF_Key[122,11]:=1854590486;
   	OWF_Key[122,12]:=1598936227;
   	OWF_Key[123,9]:=1515977147;
   	OWF_Key[123,10]:=2061812701;
   	OWF_Key[123,11]:=1866013687;
   	OWF_Key[123,12]:=4607802;
   	OWF_Key[124,9]:=810728640;
   	OWF_Key[124,10]:=768833928;
   	OWF_Key[124,11]:=1467392700;
   	OWF_Key[124,12]:=558603998;
   	OWF_Key[125,9]:=1751713093;
   	OWF_Key[125,10]:=1256264550;
   	OWF_Key[125,11]:=1970490133;
   	OWF_Key[125,12]:=1806329363;
   	OWF_Key[126,9]:=2061628321;
   	OWF_Key[126,10]:=491420936;
   	OWF_Key[126,11]:=1579649068;
   	OWF_Key[126,12]:=645775554;
   	OWF_Key[127,9]:=1507050286;
   	OWF_Key[127,10]:=47571167;
   	OWF_Key[127,11]:=1198497625;
   	OWF_Key[127,12]:=1844556864;
   	OWF_Key[128,9]:=937092274;
   	OWF_Key[128,10]:=2066941901;
   	OWF_Key[128,11]:=2088749829;
   	OWF_Key[128,12]:=1989212766;
   	OWF_Key[129,9]:=2027130018;
   	OWF_Key[129,10]:=1175951777;
   	OWF_Key[129,11]:=1971703624;
   	OWF_Key[129,12]:=1354248662;
   	OWF_Key[130,9]:=1712832844;
   	OWF_Key[130,10]:=979170224;
   	OWF_Key[130,11]:=649106733;
   	OWF_Key[130,12]:=253692714;
   	OWF_Key[131,9]:=595651429;
   	OWF_Key[131,10]:=1549613096;
   	OWF_Key[131,11]:=1452643348;
   	OWF_Key[131,12]:=58525411;
   	OWF_Key[132,9]:=997894886;
   	OWF_Key[132,10]:=1297184346;
   	OWF_Key[132,11]:=824388903;
   	OWF_Key[132,12]:=1363862442;
   	OWF_Key[133,9]:=1090176764;
   	OWF_Key[133,10]:=1282529250;
   	OWF_Key[133,11]:=1420926961;
   	OWF_Key[133,12]:=1615530204;
   	OWF_Key[134,9]:=1744742856;
   	OWF_Key[134,10]:=1213404537;
   	OWF_Key[134,11]:=1839661814;
   	OWF_Key[134,12]:=319669959;
   	OWF_Key[135,9]:=1647640650;
   	OWF_Key[135,10]:=31197237;
   	OWF_Key[135,11]:=342640965;
   	OWF_Key[135,12]:=1940913042;
   	OWF_Key[136,9]:=673587030;
   	OWF_Key[136,10]:=16922251;
   	OWF_Key[136,11]:=2016211880;
   	OWF_Key[136,12]:=284837651;
   	OWF_Key[137,9]:=1935217629;
   	OWF_Key[137,10]:=793275151;
   	OWF_Key[137,11]:=2072532760;
   	OWF_Key[137,12]:=2048048010;
   	OWF_Key[138,9]:=914987685;
   	OWF_Key[138,10]:=1965777509;
   	OWF_Key[138,11]:=2130394961;
   	OWF_Key[138,12]:=767824919;
   	OWF_Key[139,9]:=60117784;
   	OWF_Key[139,10]:=1001754166;
   	OWF_Key[139,11]:=1074350317;
   	OWF_Key[139,12]:=1528310203;
   	OWF_Key[140,9]:=108165690;
   	OWF_Key[140,10]:=1404158763;
   	OWF_Key[140,11]:=1619375742;
   	OWF_Key[140,12]:=241174143;
   	OWF_Key[141,9]:=1025074073;
   	OWF_Key[141,10]:=381400640;
   	OWF_Key[141,11]:=672604845;
   	OWF_Key[141,12]:=1687439298;
   	OWF_Key[142,9]:=405361924;
   	OWF_Key[142,10]:=1056039280;
   	OWF_Key[142,11]:=1065936229;
   	OWF_Key[142,12]:=1009892710;
   	OWF_Key[143,9]:=1397557431;
   	OWF_Key[143,10]:=1286748880;
   	OWF_Key[143,11]:=1635217434;
   	OWF_Key[143,12]:=2143552984;
   	OWF_Key[144,9]:=974809699;
   	OWF_Key[144,10]:=1030633813;
   	OWF_Key[144,11]:=914768538;
   	OWF_Key[144,12]:=988487735;
   	OWF_Key[145,9]:=1972980927;
   	OWF_Key[145,10]:=1924871894;
   	OWF_Key[145,11]:=351235414;
   	OWF_Key[145,12]:=564073825;
   	OWF_Key[146,9]:=1305901547;
   	OWF_Key[146,10]:=935924129;
   	OWF_Key[146,11]:=606118139;
   	OWF_Key[146,12]:=676806957;
   	OWF_Key[147,9]:=797894166;
   	OWF_Key[147,10]:=249563511;
   	OWF_Key[147,11]:=369911405;
   	OWF_Key[147,12]:=1718024188;
   	OWF_Key[148,9]:=445846108;
   	OWF_Key[148,10]:=1575545228;
   	OWF_Key[148,11]:=1734789187;
   	OWF_Key[148,12]:=1453154915;
   	OWF_Key[149,9]:=336541133;
   	OWF_Key[149,10]:=1892120088;
   	OWF_Key[149,11]:=808192231;
   	OWF_Key[149,12]:=2050925354;
   	OWF_Key[150,9]:=1158047330;
   	OWF_Key[150,10]:=400821636;
   	OWF_Key[150,11]:=2091245223;
   	OWF_Key[150,12]:=396677087;
   	OWF_Key[151,9]:=593738917;
   	OWF_Key[151,10]:=1819599240;
   	OWF_Key[151,11]:=528671184;
   	OWF_Key[151,12]:=1905974252;
   	OWF_Key[152,9]:=1047881867;
   	OWF_Key[152,10]:=1628041060;
   	OWF_Key[152,11]:=979770838;
   	OWF_Key[152,12]:=176104195;
   	OWF_Key[153,9]:=548455148;
   	OWF_Key[153,10]:=1899393169;
   	OWF_Key[153,11]:=364503560;
   	OWF_Key[153,12]:=1392493229;
   	OWF_Key[154,9]:=141946440;
   	OWF_Key[154,10]:=682898189;
   	OWF_Key[154,11]:=1551313638;
   	OWF_Key[154,12]:=1361870643;
   	OWF_Key[155,9]:=2007126345;
   	OWF_Key[155,10]:=1251429271;
   	OWF_Key[155,11]:=1664212479;
   	OWF_Key[155,12]:=2145730613;
   	OWF_Key[156,9]:=20326019;
   	OWF_Key[156,10]:=810173431;
   	OWF_Key[156,11]:=1519867999;
   	OWF_Key[156,12]:=1121831099;
   	OWF_Key[157,9]:=844533932;
   	OWF_Key[157,10]:=958866364;
   	OWF_Key[157,11]:=1703342512;
   	OWF_Key[157,12]:=698189185;
   	OWF_Key[158,9]:=990242471;
   	OWF_Key[158,10]:=318491994;
   	OWF_Key[158,11]:=329640992;
   	OWF_Key[158,12]:=1106957248;
   	OWF_Key[159,9]:=1980788379;
   	OWF_Key[159,10]:=886208968;
   	OWF_Key[159,11]:=1664192296;
   	OWF_Key[159,12]:=1783521060;
   	OWF_Key[160,9]:=123856352;
   	OWF_Key[160,10]:=973315151;
   	OWF_Key[160,11]:=989792177;
   	OWF_Key[160,12]:=1518147729;
   	OWF_Key[161,9]:=661702265;
   	OWF_Key[161,10]:=892864790;
   	OWF_Key[161,11]:=1819896333;
   	OWF_Key[161,12]:=453745131;
   	OWF_Key[162,9]:=1123515971;
   	OWF_Key[162,10]:=1727347230;
   	OWF_Key[162,11]:=1723323245;
   	OWF_Key[162,12]:=359175669;
   	OWF_Key[163,9]:=220624552;
   	OWF_Key[163,10]:=6972946;
   	OWF_Key[163,11]:=1837556251;
   	OWF_Key[163,12]:=433519189;
   	OWF_Key[164,9]:=385343666;
   	OWF_Key[164,10]:=445046119;
   	OWF_Key[164,11]:=344997648;
   	OWF_Key[164,12]:=927173313;
   	OWF_Key[165,9]:=277261975;
   	OWF_Key[165,10]:=1166554273;
   	OWF_Key[165,11]:=821569808;
   	OWF_Key[165,12]:=288168250;
   	OWF_Key[166,9]:=556243663;
   	OWF_Key[166,10]:=1794339253;
   	OWF_Key[166,11]:=453385726;
   	OWF_Key[166,12]:=604497673;
   	OWF_Key[167,9]:=1874617769;
   	OWF_Key[167,10]:=1319208035;
   	OWF_Key[167,11]:=504452567;
   	OWF_Key[167,12]:=1871921528;
   	OWF_Key[168,9]:=1636719299;
   	OWF_Key[168,10]:=1493960437;
   	OWF_Key[168,11]:=1254560368;
   	OWF_Key[168,12]:=1844284846;
   	OWF_Key[169,9]:=1199328367;
   	OWF_Key[169,10]:=1366035851;
   	OWF_Key[169,11]:=1209080795;
   	OWF_Key[169,12]:=629272967;
   	OWF_Key[170,9]:=1457223138;
   	OWF_Key[170,10]:=1996810357;
   	OWF_Key[170,11]:=1832711333;
   	OWF_Key[170,12]:=1314741754;
   	OWF_Key[171,9]:=1927447756;
   	OWF_Key[171,10]:=2005946028;
   	OWF_Key[171,11]:=1190514520;
   	OWF_Key[171,12]:=1363701146;
   	OWF_Key[172,9]:=704738660;
   	OWF_Key[172,10]:=651671853;
   	OWF_Key[172,11]:=348132544;
   	OWF_Key[172,12]:=2034699283;
   	OWF_Key[173,9]:=582484492;
   	OWF_Key[173,10]:=789036184;
   	OWF_Key[173,11]:=1412204677;
   	OWF_Key[173,12]:=72014072;
   	OWF_Key[174,9]:=684574399;
   	OWF_Key[174,10]:=326867321;
   	OWF_Key[174,11]:=1410824297;
   	OWF_Key[174,12]:=1593067911;
   	OWF_Key[175,9]:=73673899;
   	OWF_Key[175,10]:=1962176145;
   	OWF_Key[175,11]:=66739570;
   	OWF_Key[175,12]:=152450261;
   	OWF_Key[176,9]:=1895340919;
   	OWF_Key[176,10]:=2128297498;
   	OWF_Key[176,11]:=1815096216;
   	OWF_Key[176,12]:=591981823;
   	OWF_Key[177,9]:=1901787571;
   	OWF_Key[177,10]:=1561182749;
   	OWF_Key[177,11]:=1610342540;
   	OWF_Key[177,12]:=1354782866;
   	OWF_Key[178,9]:=56275934;
   	OWF_Key[178,10]:=1543959832;
   	OWF_Key[178,11]:=1746687655;
   	OWF_Key[178,12]:=998810497;
   	OWF_Key[179,9]:=1426969286;
   	OWF_Key[179,10]:=562521659;
   	OWF_Key[179,11]:=662837545;
   	OWF_Key[179,12]:=1705872769;
   	OWF_Key[180,9]:=206309650;
   	OWF_Key[180,10]:=1616421653;
   	OWF_Key[180,11]:=939135889;
   	OWF_Key[180,12]:=1841182941;
   	OWF_Key[181,9]:=1320846402;
   	OWF_Key[181,10]:=1280637325;
   	OWF_Key[181,11]:=873876123;
   	OWF_Key[181,12]:=1279939126;
   	OWF_Key[182,9]:=974837765;
   	OWF_Key[182,10]:=1889668126;
   	OWF_Key[182,11]:=1582978187;
   	OWF_Key[182,12]:=1306044079;
   	OWF_Key[183,9]:=905488926;
   	OWF_Key[183,10]:=897762123;
   	OWF_Key[183,11]:=1496114397;
   	OWF_Key[183,12]:=191884519;
   	OWF_Key[184,9]:=970294890;
   	OWF_Key[184,10]:=1822832783;
   	OWF_Key[184,11]:=1258160513;
   	OWF_Key[184,12]:=1424707104;
   	OWF_Key[185,9]:=849101599;
   	OWF_Key[185,10]:=1583602782;
